(* Logix 5000 project; controller FV vendor 1 type 14 code 217 rev 31.11; software revision 31.00; part 47 of 63 *)
(* tags used below, declared in another part *)
   CWD : CHECKWORD_FLAGS;
   Delphi_Does_Eng_Func : BOOL;
   FV_FV13C : PlantItem;   // FV13C
   FV_FV13J : PlantItem;   // FV13J
   FV_FV14C : PlantItem;   // FV14C
   FV_FV14J : PlantItem;   // FV14J
   FV_FV15C : PlantItem;   // FV15C
   FV_FV15J : PlantItem;   // FV15J
   FV_FV16C : PlantItem;   // FV16C
   FV_FV16J : PlantItem;   // FV16J
   FV_FV17C : PlantItem;   // FV17C
   FV_FV17J : PlantItem;   // FV17J
   FV_FV18C : PlantItem;   // FV18C
   FV_FV18J : PlantItem;   // FV18J
   FV_FV19C : PlantItem;   // FV19C
   FV_FV19J : PlantItem;   // FV19J
   FV_FV20C : PlantItem;   // FV20C
   FV_FV20J : PlantItem;   // FV20J
   FV_FV21C : PlantItem;   // FV21C
   FV_FV21J : PlantItem;   // FV21J
   FV_FV22C : PlantItem;   // FV22C
   FV_FV22J : PlantItem;   // FV22J
   FV_FV23C : PlantItem;   // FV23C
   FV_FV23J : PlantItem;   // FV23J
   FV_FV24C : PlantItem;   // FV24C
   FV_FV24J : PlantItem;   // FV24J
   FV_N255 : INT[255];   // Old Checkwords to keep Delphi working in the interim before full changeover.
(* FV_Common, continued *)

   24: [XIC(Delphi_Does_Eng_Func) [[XIC(FV_N255[25].8) [OTL(FV_FV13C.CW.[CWD.MANUAL]) ,XIC(FV_N255[25].9) OTL(FV_FV13C.CW.[CWD.MANDRV]) ,XIO(FV_N255[25].9) OTU(FV_FV13C.CW.[CWD.MANDRV]) ] ,XIO(FV_N255[25].8) [OTU(FV_FV13C.CW.[CWD.MANUAL]) ,[XIC(FV_FV13C.CW.[CWD.OUTPUT]) OTL(FV_N255[25].9) ,XIO(FV_FV13C.CW.[CWD.OUTPUT]) OTU(FV_N255[25].9) ] ] ] ,[XIC(FV_N255[25].13) OTL(FV_FV13C.CW.[CWD.CHECKOFF]) ,XIO(FV_N255[25].13) OTU(FV_FV13C.CW.[CWD.CHECKOFF]) ] ] ,XIO(Delphi_Does_Eng_Func) [[XIC(FV_FV13C.CW.[CWD.MANUAL]) OTL(FV_N255[25].8) ,XIO(FV_FV13C.CW.[CWD.MANUAL]) OTU(FV_N255[25].8) ] ,[XIC(FV_FV13C.CW.[CWD.CHECKOFF]) OTL(FV_N255[25].13) ,XIO(FV_FV13C.CW.[CWD.CHECKOFF]) OTU(FV_N255[25].13) ] ,[XIC(FV_FV13C.CW.[CWD.OUTPUT]) OTL(FV_N255[25].9) ,XIO(FV_FV13C.CW.[CWD.OUTPUT]) OTU(FV_N255[25].9) ] ] ,XIC(FV_FV13C.CW.[CWD.OUTPUT]) OTE(FV_N255[25].10) ,XIO(FV_FV13C.CW.[CWD.OUTPUT]) OTE(FV_N255[25].11) ,XIC(FV_FV13C.CW.[CWD.FAULT]) OTE(FV_N255[25].15) ];
   25: [XIC(Delphi_Does_Eng_Func) [[XIC(FV_N255[26].8) [OTL(FV_FV13J.CW.[CWD.MANUAL]) ,XIC(FV_N255[26].9) OTL(FV_FV13J.CW.[CWD.MANDRV]) ,XIO(FV_N255[26].9) OTU(FV_FV13J.CW.[CWD.MANDRV]) ] ,XIO(FV_N255[26].8) [OTU(FV_FV13J.CW.[CWD.MANUAL]) ,[XIC(FV_FV13J.CW.[CWD.OUTPUT]) OTL(FV_N255[26].9) ,XIO(FV_FV13J.CW.[CWD.OUTPUT]) OTU(FV_N255[26].9) ] ] ] ,[XIC(FV_N255[26].13) OTL(FV_FV13J.CW.[CWD.CHECKOFF]) ,XIO(FV_N255[26].13) OTU(FV_FV13J.CW.[CWD.CHECKOFF]) ] ] ,XIO(Delphi_Does_Eng_Func) [[XIC(FV_FV13J.CW.[CWD.MANUAL]) OTL(FV_N255[26].8) ,XIO(FV_FV13J.CW.[CWD.MANUAL]) OTU(FV_N255[26].8) ] ,[XIC(FV_FV13J.CW.[CWD.CHECKOFF]) OTL(FV_N255[26].13) ,XIO(FV_FV13J.CW.[CWD.CHECKOFF]) OTU(FV_N255[26].13) ] ,[XIC(FV_FV13J.CW.[CWD.OUTPUT]) OTL(FV_N255[26].9) ,XIO(FV_FV13J.CW.[CWD.OUTPUT]) OTU(FV_N255[26].9) ] ] ,XIC(FV_FV13J.CW.[CWD.OUTPUT]) OTE(FV_N255[26].10) ,XIO(FV_FV13J.CW.[CWD.OUTPUT]) OTE(FV_N255[26].11) ,XIC(FV_FV13J.CW.[CWD.FAULT]) OTE(FV_N255[26].15) ];
   26: [XIC(Delphi_Does_Eng_Func) [[XIC(FV_N255[27].8) [OTL(FV_FV14C.CW.[CWD.MANUAL]) ,XIC(FV_N255[27].9) OTL(FV_FV14C.CW.[CWD.MANDRV]) ,XIO(FV_N255[27].9) OTU(FV_FV14C.CW.[CWD.MANDRV]) ] ,XIO(FV_N255[27].8) [OTU(FV_FV14C.CW.[CWD.MANUAL]) ,[XIC(FV_FV14C.CW.[CWD.OUTPUT]) OTL(FV_N255[27].9) ,XIO(FV_FV14C.CW.[CWD.OUTPUT]) OTU(FV_N255[27].9) ] ] ] ,[XIC(FV_N255[27].13) OTL(FV_FV14C.CW.[CWD.CHECKOFF]) ,XIO(FV_N255[27].13) OTU(FV_FV14C.CW.[CWD.CHECKOFF]) ] ] ,XIO(Delphi_Does_Eng_Func) [[XIC(FV_FV14C.CW.[CWD.MANUAL]) OTL(FV_N255[27].8) ,XIO(FV_FV14C.CW.[CWD.MANUAL]) OTU(FV_N255[27].8) ] ,[XIC(FV_FV14C.CW.[CWD.CHECKOFF]) OTL(FV_N255[27].13) ,XIO(FV_FV14C.CW.[CWD.CHECKOFF]) OTU(FV_N255[27].13) ] ,[XIC(FV_FV14C.CW.[CWD.OUTPUT]) OTL(FV_N255[27].9) ,XIO(FV_FV14C.CW.[CWD.OUTPUT]) OTU(FV_N255[27].9) ] ] ,XIC(FV_FV14C.CW.[CWD.OUTPUT]) OTE(FV_N255[27].10) ,XIO(FV_FV14C.CW.[CWD.OUTPUT]) OTE(FV_N255[27].11) ,XIC(FV_FV14C.CW.[CWD.FAULT]) OTE(FV_N255[27].15) ];
   27: [XIC(Delphi_Does_Eng_Func) [[XIC(FV_N255[28].8) [OTL(FV_FV14J.CW.[CWD.MANUAL]) ,XIC(FV_N255[28].9) OTL(FV_FV14J.CW.[CWD.MANDRV]) ,XIO(FV_N255[28].9) OTU(FV_FV14J.CW.[CWD.MANDRV]) ] ,XIO(FV_N255[28].8) [OTU(FV_FV14J.CW.[CWD.MANUAL]) ,[XIC(FV_FV14J.CW.[CWD.OUTPUT]) OTL(FV_N255[28].9) ,XIO(FV_FV14J.CW.[CWD.OUTPUT]) OTU(FV_N255[28].9) ] ] ] ,[XIC(FV_N255[28].13) OTL(FV_FV14J.CW.[CWD.CHECKOFF]) ,XIO(FV_N255[28].13) OTU(FV_FV14J.CW.[CWD.CHECKOFF]) ] ] ,XIO(Delphi_Does_Eng_Func) [[XIC(FV_FV14J.CW.[CWD.MANUAL]) OTL(FV_N255[28].8) ,XIO(FV_FV14J.CW.[CWD.MANUAL]) OTU(FV_N255[28].8) ] ,[XIC(FV_FV14J.CW.[CWD.CHECKOFF]) OTL(FV_N255[28].13) ,XIO(FV_FV14J.CW.[CWD.CHECKOFF]) OTU(FV_N255[28].13) ] ,[XIC(FV_FV14J.CW.[CWD.OUTPUT]) OTL(FV_N255[28].9) ,XIO(FV_FV14J.CW.[CWD.OUTPUT]) OTU(FV_N255[28].9) ] ] ,XIC(FV_FV14J.CW.[CWD.OUTPUT]) OTE(FV_N255[28].10) ,XIO(FV_FV14J.CW.[CWD.OUTPUT]) OTE(FV_N255[28].11) ,XIC(FV_FV14J.CW.[CWD.FAULT]) OTE(FV_N255[28].15) ];
   28: [XIC(Delphi_Does_Eng_Func) [[XIC(FV_N255[29].8) [OTL(FV_FV15C.CW.[CWD.MANUAL]) ,XIC(FV_N255[29].9) OTL(FV_FV15C.CW.[CWD.MANDRV]) ,XIO(FV_N255[29].9) OTU(FV_FV15C.CW.[CWD.MANDRV]) ] ,XIO(FV_N255[29].8) [OTU(FV_FV15C.CW.[CWD.MANUAL]) ,[XIC(FV_FV15C.CW.[CWD.OUTPUT]) OTL(FV_N255[29].9) ,XIO(FV_FV15C.CW.[CWD.OUTPUT]) OTU(FV_N255[29].9) ] ] ] ,[XIC(FV_N255[29].13) OTL(FV_FV15C.CW.[CWD.CHECKOFF]) ,XIO(FV_N255[29].13) OTU(FV_FV15C.CW.[CWD.CHECKOFF]) ] ] ,XIO(Delphi_Does_Eng_Func) [[XIC(FV_FV15C.CW.[CWD.MANUAL]) OTL(FV_N255[29].8) ,XIO(FV_FV15C.CW.[CWD.MANUAL]) OTU(FV_N255[29].8) ] ,[XIC(FV_FV15C.CW.[CWD.CHECKOFF]) OTL(FV_N255[29].13) ,XIO(FV_FV15C.CW.[CWD.CHECKOFF]) OTU(FV_N255[29].13) ] ,[XIC(FV_FV15C.CW.[CWD.OUTPUT]) OTL(FV_N255[29].9) ,XIO(FV_FV15C.CW.[CWD.OUTPUT]) OTU(FV_N255[29].9) ] ] ,XIC(FV_FV15C.CW.[CWD.OUTPUT]) OTE(FV_N255[29].10) ,XIO(FV_FV15C.CW.[CWD.OUTPUT]) OTE(FV_N255[29].11) ,XIC(FV_FV15C.CW.[CWD.FAULT]) OTE(FV_N255[29].15) ];
   29: [XIC(Delphi_Does_Eng_Func) [[XIC(FV_N255[30].8) [OTL(FV_FV15J.CW.[CWD.MANUAL]) ,XIC(FV_N255[30].9) OTL(FV_FV15J.CW.[CWD.MANDRV]) ,XIO(FV_N255[30].9) OTU(FV_FV15J.CW.[CWD.MANDRV]) ] ,XIO(FV_N255[30].8) [OTU(FV_FV15J.CW.[CWD.MANUAL]) ,[XIC(FV_FV15J.CW.[CWD.OUTPUT]) OTL(FV_N255[30].9) ,XIO(FV_FV15J.CW.[CWD.OUTPUT]) OTU(FV_N255[30].9) ] ] ] ,[XIC(FV_N255[30].13) OTL(FV_FV15J.CW.[CWD.CHECKOFF]) ,XIO(FV_N255[30].13) OTU(FV_FV15J.CW.[CWD.CHECKOFF]) ] ] ,XIO(Delphi_Does_Eng_Func) [[XIC(FV_FV15J.CW.[CWD.MANUAL]) OTL(FV_N255[30].8) ,XIO(FV_FV15J.CW.[CWD.MANUAL]) OTU(FV_N255[30].8) ] ,[XIC(FV_FV15J.CW.[CWD.CHECKOFF]) OTL(FV_N255[30].13) ,XIO(FV_FV15J.CW.[CWD.CHECKOFF]) OTU(FV_N255[30].13) ] ,[XIC(FV_FV15J.CW.[CWD.OUTPUT]) OTL(FV_N255[30].9) ,XIO(FV_FV15J.CW.[CWD.OUTPUT]) OTU(FV_N255[30].9) ] ] ,XIC(FV_FV15J.CW.[CWD.OUTPUT]) OTE(FV_N255[30].10) ,XIO(FV_FV15J.CW.[CWD.OUTPUT]) OTE(FV_N255[30].11) ,XIC(FV_FV15J.CW.[CWD.FAULT]) OTE(FV_N255[30].15) ];
   30: [XIC(Delphi_Does_Eng_Func) [[XIC(FV_N255[31].8) [OTL(FV_FV16C.CW.[CWD.MANUAL]) ,XIC(FV_N255[31].9) OTL(FV_FV16C.CW.[CWD.MANDRV]) ,XIO(FV_N255[31].9) OTU(FV_FV16C.CW.[CWD.MANDRV]) ] ,XIO(FV_N255[31].8) [OTU(FV_FV16C.CW.[CWD.MANUAL]) ,[XIC(FV_FV16C.CW.[CWD.OUTPUT]) OTL(FV_N255[31].9) ,XIO(FV_FV16C.CW.[CWD.OUTPUT]) OTU(FV_N255[31].9) ] ] ] ,[XIC(FV_N255[31].13) OTL(FV_FV16C.CW.[CWD.CHECKOFF]) ,XIO(FV_N255[31].13) OTU(FV_FV16C.CW.[CWD.CHECKOFF]) ] ] ,XIO(Delphi_Does_Eng_Func) [[XIC(FV_FV16C.CW.[CWD.MANUAL]) OTL(FV_N255[31].8) ,XIO(FV_FV16C.CW.[CWD.MANUAL]) OTU(FV_N255[31].8) ] ,[XIC(FV_FV16C.CW.[CWD.CHECKOFF]) OTL(FV_N255[31].13) ,XIO(FV_FV16C.CW.[CWD.CHECKOFF]) OTU(FV_N255[31].13) ] ,[XIC(FV_FV16C.CW.[CWD.OUTPUT]) OTL(FV_N255[31].9) ,XIO(FV_FV16C.CW.[CWD.OUTPUT]) OTU(FV_N255[31].9) ] ] ,XIC(FV_FV16C.CW.[CWD.OUTPUT]) OTE(FV_N255[31].10) ,XIO(FV_FV16C.CW.[CWD.OUTPUT]) OTE(FV_N255[31].11) ,XIC(FV_FV16C.CW.[CWD.FAULT]) OTE(FV_N255[31].15) ];
   31: [XIC(Delphi_Does_Eng_Func) [[XIC(FV_N255[32].8) [OTL(FV_FV16J.CW.[CWD.MANUAL]) ,XIC(FV_N255[32].9) OTL(FV_FV16J.CW.[CWD.MANDRV]) ,XIO(FV_N255[32].9) OTU(FV_FV16J.CW.[CWD.MANDRV]) ] ,XIO(FV_N255[32].8) [OTU(FV_FV16J.CW.[CWD.MANUAL]) ,[XIC(FV_FV16J.CW.[CWD.OUTPUT]) OTL(FV_N255[32].9) ,XIO(FV_FV16J.CW.[CWD.OUTPUT]) OTU(FV_N255[32].9) ] ] ] ,[XIC(FV_N255[32].13) OTL(FV_FV16J.CW.[CWD.CHECKOFF]) ,XIO(FV_N255[32].13) OTU(FV_FV16J.CW.[CWD.CHECKOFF]) ] ] ,XIO(Delphi_Does_Eng_Func) [[XIC(FV_FV16J.CW.[CWD.MANUAL]) OTL(FV_N255[32].8) ,XIO(FV_FV16J.CW.[CWD.MANUAL]) OTU(FV_N255[32].8) ] ,[XIC(FV_FV16J.CW.[CWD.CHECKOFF]) OTL(FV_N255[32].13) ,XIO(FV_FV16J.CW.[CWD.CHECKOFF]) OTU(FV_N255[32].13) ] ,[XIC(FV_FV16J.CW.[CWD.OUTPUT]) OTL(FV_N255[32].9) ,XIO(FV_FV16J.CW.[CWD.OUTPUT]) OTU(FV_N255[32].9) ] ] ,XIC(FV_FV16J.CW.[CWD.OUTPUT]) OTE(FV_N255[32].10) ,XIO(FV_FV16J.CW.[CWD.OUTPUT]) OTE(FV_N255[32].11) ,XIC(FV_FV16J.CW.[CWD.FAULT]) OTE(FV_N255[32].15) ];
   32: [XIC(Delphi_Does_Eng_Func) [[XIC(FV_N255[33].8) [OTL(FV_FV17C.CW.[CWD.MANUAL]) ,XIC(FV_N255[33].9) OTL(FV_FV17C.CW.[CWD.MANDRV]) ,XIO(FV_N255[33].9) OTU(FV_FV17C.CW.[CWD.MANDRV]) ] ,XIO(FV_N255[33].8) [OTU(FV_FV17C.CW.[CWD.MANUAL]) ,[XIC(FV_FV17C.CW.[CWD.OUTPUT]) OTL(FV_N255[33].9) ,XIO(FV_FV17C.CW.[CWD.OUTPUT]) OTU(FV_N255[33].9) ] ] ] ,[XIC(FV_N255[33].13) OTL(FV_FV17C.CW.[CWD.CHECKOFF]) ,XIO(FV_N255[33].13) OTU(FV_FV17C.CW.[CWD.CHECKOFF]) ] ] ,XIO(Delphi_Does_Eng_Func) [[XIC(FV_FV17C.CW.[CWD.MANUAL]) OTL(FV_N255[33].8) ,XIO(FV_FV17C.CW.[CWD.MANUAL]) OTU(FV_N255[33].8) ] ,[XIC(FV_FV17C.CW.[CWD.CHECKOFF]) OTL(FV_N255[33].13) ,XIO(FV_FV17C.CW.[CWD.CHECKOFF]) OTU(FV_N255[33].13) ] ,[XIC(FV_FV17C.CW.[CWD.OUTPUT]) OTL(FV_N255[33].9) ,XIO(FV_FV17C.CW.[CWD.OUTPUT]) OTU(FV_N255[33].9) ] ] ,XIC(FV_FV17C.CW.[CWD.OUTPUT]) OTE(FV_N255[33].10) ,XIO(FV_FV17C.CW.[CWD.OUTPUT]) OTE(FV_N255[33].11) ,XIC(FV_FV17C.CW.[CWD.FAULT]) OTE(FV_N255[33].15) ];
   33: [XIC(Delphi_Does_Eng_Func) [[XIC(FV_N255[34].8) [OTL(FV_FV17J.CW.[CWD.MANUAL]) ,XIC(FV_N255[34].9) OTL(FV_FV17J.CW.[CWD.MANDRV]) ,XIO(FV_N255[34].9) OTU(FV_FV17J.CW.[CWD.MANDRV]) ] ,XIO(FV_N255[34].8) [OTU(FV_FV17J.CW.[CWD.MANUAL]) ,[XIC(FV_FV17J.CW.[CWD.OUTPUT]) OTL(FV_N255[34].9) ,XIO(FV_FV17J.CW.[CWD.OUTPUT]) OTU(FV_N255[34].9) ] ] ] ,[XIC(FV_N255[34].13) OTL(FV_FV17J.CW.[CWD.CHECKOFF]) ,XIO(FV_N255[34].13) OTU(FV_FV17J.CW.[CWD.CHECKOFF]) ] ] ,XIO(Delphi_Does_Eng_Func) [[XIC(FV_FV17J.CW.[CWD.MANUAL]) OTL(FV_N255[34].8) ,XIO(FV_FV17J.CW.[CWD.MANUAL]) OTU(FV_N255[34].8) ] ,[XIC(FV_FV17J.CW.[CWD.CHECKOFF]) OTL(FV_N255[34].13) ,XIO(FV_FV17J.CW.[CWD.CHECKOFF]) OTU(FV_N255[34].13) ] ,[XIC(FV_FV17J.CW.[CWD.OUTPUT]) OTL(FV_N255[34].9) ,XIO(FV_FV17J.CW.[CWD.OUTPUT]) OTU(FV_N255[34].9) ] ] ,XIC(FV_FV17J.CW.[CWD.OUTPUT]) OTE(FV_N255[34].10) ,XIO(FV_FV17J.CW.[CWD.OUTPUT]) OTE(FV_N255[34].11) ,XIC(FV_FV17J.CW.[CWD.FAULT]) OTE(FV_N255[34].15) ];
   34: [XIC(Delphi_Does_Eng_Func) [[XIC(FV_N255[35].8) [OTL(FV_FV18C.CW.[CWD.MANUAL]) ,XIC(FV_N255[35].9) OTL(FV_FV18C.CW.[CWD.MANDRV]) ,XIO(FV_N255[35].9) OTU(FV_FV18C.CW.[CWD.MANDRV]) ] ,XIO(FV_N255[35].8) [OTU(FV_FV18C.CW.[CWD.MANUAL]) ,[XIC(FV_FV18C.CW.[CWD.OUTPUT]) OTL(FV_N255[35].9) ,XIO(FV_FV18C.CW.[CWD.OUTPUT]) OTU(FV_N255[35].9) ] ] ] ,[XIC(FV_N255[35].13) OTL(FV_FV18C.CW.[CWD.CHECKOFF]) ,XIO(FV_N255[35].13) OTU(FV_FV18C.CW.[CWD.CHECKOFF]) ] ] ,XIO(Delphi_Does_Eng_Func) [[XIC(FV_FV18C.CW.[CWD.MANUAL]) OTL(FV_N255[35].8) ,XIO(FV_FV18C.CW.[CWD.MANUAL]) OTU(FV_N255[35].8) ] ,[XIC(FV_FV18C.CW.[CWD.CHECKOFF]) OTL(FV_N255[35].13) ,XIO(FV_FV18C.CW.[CWD.CHECKOFF]) OTU(FV_N255[35].13) ] ,[XIC(FV_FV18C.CW.[CWD.OUTPUT]) OTL(FV_N255[35].9) ,XIO(FV_FV18C.CW.[CWD.OUTPUT]) OTU(FV_N255[35].9) ] ] ,XIC(FV_FV18C.CW.[CWD.OUTPUT]) OTE(FV_N255[35].10) ,XIO(FV_FV18C.CW.[CWD.OUTPUT]) OTE(FV_N255[35].11) ,XIC(FV_FV18C.CW.[CWD.FAULT]) OTE(FV_N255[35].15) ];
   35: [XIC(Delphi_Does_Eng_Func) [[XIC(FV_N255[36].8) [OTL(FV_FV18J.CW.[CWD.MANUAL]) ,XIC(FV_N255[36].9) OTL(FV_FV18J.CW.[CWD.MANDRV]) ,XIO(FV_N255[36].9) OTU(FV_FV18J.CW.[CWD.MANDRV]) ] ,XIO(FV_N255[36].8) [OTU(FV_FV18J.CW.[CWD.MANUAL]) ,[XIC(FV_FV18J.CW.[CWD.OUTPUT]) OTL(FV_N255[36].9) ,XIO(FV_FV18J.CW.[CWD.OUTPUT]) OTU(FV_N255[36].9) ] ] ] ,[XIC(FV_N255[36].13) OTL(FV_FV18J.CW.[CWD.CHECKOFF]) ,XIO(FV_N255[36].13) OTU(FV_FV18J.CW.[CWD.CHECKOFF]) ] ] ,XIO(Delphi_Does_Eng_Func) [[XIC(FV_FV18J.CW.[CWD.MANUAL]) OTL(FV_N255[36].8) ,XIO(FV_FV18J.CW.[CWD.MANUAL]) OTU(FV_N255[36].8) ] ,[XIC(FV_FV18J.CW.[CWD.CHECKOFF]) OTL(FV_N255[36].13) ,XIO(FV_FV18J.CW.[CWD.CHECKOFF]) OTU(FV_N255[36].13) ] ,[XIC(FV_FV18J.CW.[CWD.OUTPUT]) OTL(FV_N255[36].9) ,XIO(FV_FV18J.CW.[CWD.OUTPUT]) OTU(FV_N255[36].9) ] ] ,XIC(FV_FV18J.CW.[CWD.OUTPUT]) OTE(FV_N255[36].10) ,XIO(FV_FV18J.CW.[CWD.OUTPUT]) OTE(FV_N255[36].11) ,XIC(FV_FV18J.CW.[CWD.FAULT]) OTE(FV_N255[36].15) ];
   36: [XIC(Delphi_Does_Eng_Func) [[XIC(FV_N255[37].8) [OTL(FV_FV19C.CW.[CWD.MANUAL]) ,XIC(FV_N255[37].9) OTL(FV_FV19C.CW.[CWD.MANDRV]) ,XIO(FV_N255[37].9) OTU(FV_FV19C.CW.[CWD.MANDRV]) ] ,XIO(FV_N255[37].8) [OTU(FV_FV19C.CW.[CWD.MANUAL]) ,[XIC(FV_FV19C.CW.[CWD.OUTPUT]) OTL(FV_N255[37].9) ,XIO(FV_FV19C.CW.[CWD.OUTPUT]) OTU(FV_N255[37].9) ] ] ] ,[XIC(FV_N255[37].13) OTL(FV_FV19C.CW.[CWD.CHECKOFF]) ,XIO(FV_N255[37].13) OTU(FV_FV19C.CW.[CWD.CHECKOFF]) ] ] ,XIO(Delphi_Does_Eng_Func) [[XIC(FV_FV19C.CW.[CWD.MANUAL]) OTL(FV_N255[37].8) ,XIO(FV_FV19C.CW.[CWD.MANUAL]) OTU(FV_N255[37].8) ] ,[XIC(FV_FV19C.CW.[CWD.CHECKOFF]) OTL(FV_N255[37].13) ,XIO(FV_FV19C.CW.[CWD.CHECKOFF]) OTU(FV_N255[37].13) ] ,[XIC(FV_FV19C.CW.[CWD.OUTPUT]) OTL(FV_N255[37].9) ,XIO(FV_FV19C.CW.[CWD.OUTPUT]) OTU(FV_N255[37].9) ] ] ,XIC(FV_FV19C.CW.[CWD.OUTPUT]) OTE(FV_N255[37].10) ,XIO(FV_FV19C.CW.[CWD.OUTPUT]) OTE(FV_N255[37].11) ,XIC(FV_FV19C.CW.[CWD.FAULT]) OTE(FV_N255[37].15) ];
   37: [XIC(Delphi_Does_Eng_Func) [[XIC(FV_N255[38].8) [OTL(FV_FV19J.CW.[CWD.MANUAL]) ,XIC(FV_N255[38].9) OTL(FV_FV19J.CW.[CWD.MANDRV]) ,XIO(FV_N255[38].9) OTU(FV_FV19J.CW.[CWD.MANDRV]) ] ,XIO(FV_N255[38].8) [OTU(FV_FV19J.CW.[CWD.MANUAL]) ,[XIC(FV_FV19J.CW.[CWD.OUTPUT]) OTL(FV_N255[38].9) ,XIO(FV_FV19J.CW.[CWD.OUTPUT]) OTU(FV_N255[38].9) ] ] ] ,[XIC(FV_N255[38].13) OTL(FV_FV19J.CW.[CWD.CHECKOFF]) ,XIO(FV_N255[38].13) OTU(FV_FV19J.CW.[CWD.CHECKOFF]) ] ] ,XIO(Delphi_Does_Eng_Func) [[XIC(FV_FV19J.CW.[CWD.MANUAL]) OTL(FV_N255[38].8) ,XIO(FV_FV19J.CW.[CWD.MANUAL]) OTU(FV_N255[38].8) ] ,[XIC(FV_FV19J.CW.[CWD.CHECKOFF]) OTL(FV_N255[38].13) ,XIO(FV_FV19J.CW.[CWD.CHECKOFF]) OTU(FV_N255[38].13) ] ,[XIC(FV_FV19J.CW.[CWD.OUTPUT]) OTL(FV_N255[38].9) ,XIO(FV_FV19J.CW.[CWD.OUTPUT]) OTU(FV_N255[38].9) ] ] ,XIC(FV_FV19J.CW.[CWD.OUTPUT]) OTE(FV_N255[38].10) ,XIO(FV_FV19J.CW.[CWD.OUTPUT]) OTE(FV_N255[38].11) ,XIC(FV_FV19J.CW.[CWD.FAULT]) OTE(FV_N255[38].15) ];
   38: [XIC(Delphi_Does_Eng_Func) [[XIC(FV_N255[39].8) [OTL(FV_FV20C.CW.[CWD.MANUAL]) ,XIC(FV_N255[39].9) OTL(FV_FV20C.CW.[CWD.MANDRV]) ,XIO(FV_N255[39].9) OTU(FV_FV20C.CW.[CWD.MANDRV]) ] ,XIO(FV_N255[39].8) [OTU(FV_FV20C.CW.[CWD.MANUAL]) ,[XIC(FV_FV20C.CW.[CWD.OUTPUT]) OTL(FV_N255[39].9) ,XIO(FV_FV20C.CW.[CWD.OUTPUT]) OTU(FV_N255[39].9) ] ] ] ,[XIC(FV_N255[39].13) OTL(FV_FV20C.CW.[CWD.CHECKOFF]) ,XIO(FV_N255[39].13) OTU(FV_FV20C.CW.[CWD.CHECKOFF]) ] ] ,XIO(Delphi_Does_Eng_Func) [[XIC(FV_FV20C.CW.[CWD.MANUAL]) OTL(FV_N255[39].8) ,XIO(FV_FV20C.CW.[CWD.MANUAL]) OTU(FV_N255[39].8) ] ,[XIC(FV_FV20C.CW.[CWD.CHECKOFF]) OTL(FV_N255[39].13) ,XIO(FV_FV20C.CW.[CWD.CHECKOFF]) OTU(FV_N255[39].13) ] ,[XIC(FV_FV20C.CW.[CWD.OUTPUT]) OTL(FV_N255[39].9) ,XIO(FV_FV20C.CW.[CWD.OUTPUT]) OTU(FV_N255[39].9) ] ] ,XIC(FV_FV20C.CW.[CWD.OUTPUT]) OTE(FV_N255[39].10) ,XIO(FV_FV20C.CW.[CWD.OUTPUT]) OTE(FV_N255[39].11) ,XIC(FV_FV20C.CW.[CWD.FAULT]) OTE(FV_N255[39].15) ];
   39: [XIC(Delphi_Does_Eng_Func) [[XIC(FV_N255[40].8) [OTL(FV_FV20J.CW.[CWD.MANUAL]) ,XIC(FV_N255[40].9) OTL(FV_FV20J.CW.[CWD.MANDRV]) ,XIO(FV_N255[40].9) OTU(FV_FV20J.CW.[CWD.MANDRV]) ] ,XIO(FV_N255[40].8) [OTU(FV_FV20J.CW.[CWD.MANUAL]) ,[XIC(FV_FV20J.CW.[CWD.OUTPUT]) OTL(FV_N255[40].9) ,XIO(FV_FV20J.CW.[CWD.OUTPUT]) OTU(FV_N255[40].9) ] ] ] ,[XIC(FV_N255[40].13) OTL(FV_FV20J.CW.[CWD.CHECKOFF]) ,XIO(FV_N255[40].13) OTU(FV_FV20J.CW.[CWD.CHECKOFF]) ] ] ,XIO(Delphi_Does_Eng_Func) [[XIC(FV_FV20J.CW.[CWD.MANUAL]) OTL(FV_N255[40].8) ,XIO(FV_FV20J.CW.[CWD.MANUAL]) OTU(FV_N255[40].8) ] ,[XIC(FV_FV20J.CW.[CWD.CHECKOFF]) OTL(FV_N255[40].13) ,XIO(FV_FV20J.CW.[CWD.CHECKOFF]) OTU(FV_N255[40].13) ] ,[XIC(FV_FV20J.CW.[CWD.OUTPUT]) OTL(FV_N255[40].9) ,XIO(FV_FV20J.CW.[CWD.OUTPUT]) OTU(FV_N255[40].9) ] ] ,XIC(FV_FV20J.CW.[CWD.OUTPUT]) OTE(FV_N255[40].10) ,XIO(FV_FV20J.CW.[CWD.OUTPUT]) OTE(FV_N255[40].11) ,XIC(FV_FV20J.CW.[CWD.FAULT]) OTE(FV_N255[40].15) ];
   40: [XIC(Delphi_Does_Eng_Func) [[XIC(FV_N255[41].8) [OTL(FV_FV21C.CW.[CWD.MANUAL]) ,XIC(FV_N255[41].9) OTL(FV_FV21C.CW.[CWD.MANDRV]) ,XIO(FV_N255[41].9) OTU(FV_FV21C.CW.[CWD.MANDRV]) ] ,XIO(FV_N255[41].8) [OTU(FV_FV21C.CW.[CWD.MANUAL]) ,[XIC(FV_FV21C.CW.[CWD.OUTPUT]) OTL(FV_N255[41].9) ,XIO(FV_FV21C.CW.[CWD.OUTPUT]) OTU(FV_N255[41].9) ] ] ] ,[XIC(FV_N255[41].13) OTL(FV_FV21C.CW.[CWD.CHECKOFF]) ,XIO(FV_N255[41].13) OTU(FV_FV21C.CW.[CWD.CHECKOFF]) ] ] ,XIO(Delphi_Does_Eng_Func) [[XIC(FV_FV21C.CW.[CWD.MANUAL]) OTL(FV_N255[41].8) ,XIO(FV_FV21C.CW.[CWD.MANUAL]) OTU(FV_N255[41].8) ] ,[XIC(FV_FV21C.CW.[CWD.CHECKOFF]) OTL(FV_N255[41].13) ,XIO(FV_FV21C.CW.[CWD.CHECKOFF]) OTU(FV_N255[41].13) ] ,[XIC(FV_FV21C.CW.[CWD.OUTPUT]) OTL(FV_N255[41].9) ,XIO(FV_FV21C.CW.[CWD.OUTPUT]) OTU(FV_N255[41].9) ] ] ,XIC(FV_FV21C.CW.[CWD.OUTPUT]) OTE(FV_N255[41].10) ,XIO(FV_FV21C.CW.[CWD.OUTPUT]) OTE(FV_N255[41].11) ,XIC(FV_FV21C.CW.[CWD.FAULT]) OTE(FV_N255[41].15) ];
   41: [XIC(Delphi_Does_Eng_Func) [[XIC(FV_N255[42].8) [OTL(FV_FV21J.CW.[CWD.MANUAL]) ,XIC(FV_N255[42].9) OTL(FV_FV21J.CW.[CWD.MANDRV]) ,XIO(FV_N255[42].9) OTU(FV_FV21J.CW.[CWD.MANDRV]) ] ,XIO(FV_N255[42].8) [OTU(FV_FV21J.CW.[CWD.MANUAL]) ,[XIC(FV_FV21J.CW.[CWD.OUTPUT]) OTL(FV_N255[42].9) ,XIO(FV_FV21J.CW.[CWD.OUTPUT]) OTU(FV_N255[42].9) ] ] ] ,[XIC(FV_N255[42].13) OTL(FV_FV21J.CW.[CWD.CHECKOFF]) ,XIO(FV_N255[42].13) OTU(FV_FV21J.CW.[CWD.CHECKOFF]) ] ] ,XIO(Delphi_Does_Eng_Func) [[XIC(FV_FV21J.CW.[CWD.MANUAL]) OTL(FV_N255[42].8) ,XIO(FV_FV21J.CW.[CWD.MANUAL]) OTU(FV_N255[42].8) ] ,[XIC(FV_FV21J.CW.[CWD.CHECKOFF]) OTL(FV_N255[42].13) ,XIO(FV_FV21J.CW.[CWD.CHECKOFF]) OTU(FV_N255[42].13) ] ,[XIC(FV_FV21J.CW.[CWD.OUTPUT]) OTL(FV_N255[42].9) ,XIO(FV_FV21J.CW.[CWD.OUTPUT]) OTU(FV_N255[42].9) ] ] ,XIC(FV_FV21J.CW.[CWD.OUTPUT]) OTE(FV_N255[42].10) ,XIO(FV_FV21J.CW.[CWD.OUTPUT]) OTE(FV_N255[42].11) ,XIC(FV_FV21J.CW.[CWD.FAULT]) OTE(FV_N255[42].15) ];
   42: [XIC(Delphi_Does_Eng_Func) [[XIC(FV_N255[43].8) [OTL(FV_FV22C.CW.[CWD.MANUAL]) ,XIC(FV_N255[43].9) OTL(FV_FV22C.CW.[CWD.MANDRV]) ,XIO(FV_N255[43].9) OTU(FV_FV22C.CW.[CWD.MANDRV]) ] ,XIO(FV_N255[43].8) [OTU(FV_FV22C.CW.[CWD.MANUAL]) ,[XIC(FV_FV22C.CW.[CWD.OUTPUT]) OTL(FV_N255[43].9) ,XIO(FV_FV22C.CW.[CWD.OUTPUT]) OTU(FV_N255[43].9) ] ] ] ,[XIC(FV_N255[43].13) OTL(FV_FV22C.CW.[CWD.CHECKOFF]) ,XIO(FV_N255[43].13) OTU(FV_FV22C.CW.[CWD.CHECKOFF]) ] ] ,XIO(Delphi_Does_Eng_Func) [[XIC(FV_FV22C.CW.[CWD.MANUAL]) OTL(FV_N255[43].8) ,XIO(FV_FV22C.CW.[CWD.MANUAL]) OTU(FV_N255[43].8) ] ,[XIC(FV_FV22C.CW.[CWD.CHECKOFF]) OTL(FV_N255[43].13) ,XIO(FV_FV22C.CW.[CWD.CHECKOFF]) OTU(FV_N255[43].13) ] ,[XIC(FV_FV22C.CW.[CWD.OUTPUT]) OTL(FV_N255[43].9) ,XIO(FV_FV22C.CW.[CWD.OUTPUT]) OTU(FV_N255[43].9) ] ] ,XIC(FV_FV22C.CW.[CWD.OUTPUT]) OTE(FV_N255[43].10) ,XIO(FV_FV22C.CW.[CWD.OUTPUT]) OTE(FV_N255[43].11) ,XIC(FV_FV22C.CW.[CWD.FAULT]) OTE(FV_N255[43].15) ];
   43: [XIC(Delphi_Does_Eng_Func) [[XIC(FV_N255[44].8) [OTL(FV_FV22J.CW.[CWD.MANUAL]) ,XIC(FV_N255[44].9) OTL(FV_FV22J.CW.[CWD.MANDRV]) ,XIO(FV_N255[44].9) OTU(FV_FV22J.CW.[CWD.MANDRV]) ] ,XIO(FV_N255[44].8) [OTU(FV_FV22J.CW.[CWD.MANUAL]) ,[XIC(FV_FV22J.CW.[CWD.OUTPUT]) OTL(FV_N255[44].9) ,XIO(FV_FV22J.CW.[CWD.OUTPUT]) OTU(FV_N255[44].9) ] ] ] ,[XIC(FV_N255[44].13) OTL(FV_FV22J.CW.[CWD.CHECKOFF]) ,XIO(FV_N255[44].13) OTU(FV_FV22J.CW.[CWD.CHECKOFF]) ] ] ,XIO(Delphi_Does_Eng_Func) [[XIC(FV_FV22J.CW.[CWD.MANUAL]) OTL(FV_N255[44].8) ,XIO(FV_FV22J.CW.[CWD.MANUAL]) OTU(FV_N255[44].8) ] ,[XIC(FV_FV22J.CW.[CWD.CHECKOFF]) OTL(FV_N255[44].13) ,XIO(FV_FV22J.CW.[CWD.CHECKOFF]) OTU(FV_N255[44].13) ] ,[XIC(FV_FV22J.CW.[CWD.OUTPUT]) OTL(FV_N255[44].9) ,XIO(FV_FV22J.CW.[CWD.OUTPUT]) OTU(FV_N255[44].9) ] ] ,XIC(FV_FV22J.CW.[CWD.OUTPUT]) OTE(FV_N255[44].10) ,XIO(FV_FV22J.CW.[CWD.OUTPUT]) OTE(FV_N255[44].11) ,XIC(FV_FV22J.CW.[CWD.FAULT]) OTE(FV_N255[44].15) ];
   44: [XIC(Delphi_Does_Eng_Func) [[XIC(FV_N255[45].8) [OTL(FV_FV23C.CW.[CWD.MANUAL]) ,XIC(FV_N255[45].9) OTL(FV_FV23C.CW.[CWD.MANDRV]) ,XIO(FV_N255[45].9) OTU(FV_FV23C.CW.[CWD.MANDRV]) ] ,XIO(FV_N255[45].8) [OTU(FV_FV23C.CW.[CWD.MANUAL]) ,[XIC(FV_FV23C.CW.[CWD.OUTPUT]) OTL(FV_N255[45].9) ,XIO(FV_FV23C.CW.[CWD.OUTPUT]) OTU(FV_N255[45].9) ] ] ] ,[XIC(FV_N255[45].13) OTL(FV_FV23C.CW.[CWD.CHECKOFF]) ,XIO(FV_N255[45].13) OTU(FV_FV23C.CW.[CWD.CHECKOFF]) ] ] ,XIO(Delphi_Does_Eng_Func) [[XIC(FV_FV23C.CW.[CWD.MANUAL]) OTL(FV_N255[45].8) ,XIO(FV_FV23C.CW.[CWD.MANUAL]) OTU(FV_N255[45].8) ] ,[XIC(FV_FV23C.CW.[CWD.CHECKOFF]) OTL(FV_N255[45].13) ,XIO(FV_FV23C.CW.[CWD.CHECKOFF]) OTU(FV_N255[45].13) ] ,[XIC(FV_FV23C.CW.[CWD.OUTPUT]) OTL(FV_N255[45].9) ,XIO(FV_FV23C.CW.[CWD.OUTPUT]) OTU(FV_N255[45].9) ] ] ,XIC(FV_FV23C.CW.[CWD.OUTPUT]) OTE(FV_N255[45].10) ,XIO(FV_FV23C.CW.[CWD.OUTPUT]) OTE(FV_N255[45].11) ,XIC(FV_FV23C.CW.[CWD.FAULT]) OTE(FV_N255[45].15) ];
   45: [XIC(Delphi_Does_Eng_Func) [[XIC(FV_N255[46].8) [OTL(FV_FV23J.CW.[CWD.MANUAL]) ,XIC(FV_N255[46].9) OTL(FV_FV23J.CW.[CWD.MANDRV]) ,XIO(FV_N255[46].9) OTU(FV_FV23J.CW.[CWD.MANDRV]) ] ,XIO(FV_N255[46].8) [OTU(FV_FV23J.CW.[CWD.MANUAL]) ,[XIC(FV_FV23J.CW.[CWD.OUTPUT]) OTL(FV_N255[46].9) ,XIO(FV_FV23J.CW.[CWD.OUTPUT]) OTU(FV_N255[46].9) ] ] ] ,[XIC(FV_N255[46].13) OTL(FV_FV23J.CW.[CWD.CHECKOFF]) ,XIO(FV_N255[46].13) OTU(FV_FV23J.CW.[CWD.CHECKOFF]) ] ] ,XIO(Delphi_Does_Eng_Func) [[XIC(FV_FV23J.CW.[CWD.MANUAL]) OTL(FV_N255[46].8) ,XIO(FV_FV23J.CW.[CWD.MANUAL]) OTU(FV_N255[46].8) ] ,[XIC(FV_FV23J.CW.[CWD.CHECKOFF]) OTL(FV_N255[46].13) ,XIO(FV_FV23J.CW.[CWD.CHECKOFF]) OTU(FV_N255[46].13) ] ,[XIC(FV_FV23J.CW.[CWD.OUTPUT]) OTL(FV_N255[46].9) ,XIO(FV_FV23J.CW.[CWD.OUTPUT]) OTU(FV_N255[46].9) ] ] ,XIC(FV_FV23J.CW.[CWD.OUTPUT]) OTE(FV_N255[46].10) ,XIO(FV_FV23J.CW.[CWD.OUTPUT]) OTE(FV_N255[46].11) ,XIC(FV_FV23J.CW.[CWD.FAULT]) OTE(FV_N255[46].15) ];
   46: [XIC(Delphi_Does_Eng_Func) [[XIC(FV_N255[47].8) [OTL(FV_FV24C.CW.[CWD.MANUAL]) ,XIC(FV_N255[47].9) OTL(FV_FV24C.CW.[CWD.MANDRV]) ,XIO(FV_N255[47].9) OTU(FV_FV24C.CW.[CWD.MANDRV]) ] ,XIO(FV_N255[47].8) [OTU(FV_FV24C.CW.[CWD.MANUAL]) ,[XIC(FV_FV24C.CW.[CWD.OUTPUT]) OTL(FV_N255[47].9) ,XIO(FV_FV24C.CW.[CWD.OUTPUT]) OTU(FV_N255[47].9) ] ] ] ,[XIC(FV_N255[47].13) OTL(FV_FV24C.CW.[CWD.CHECKOFF]) ,XIO(FV_N255[47].13) OTU(FV_FV24C.CW.[CWD.CHECKOFF]) ] ] ,XIO(Delphi_Does_Eng_Func) [[XIC(FV_FV24C.CW.[CWD.MANUAL]) OTL(FV_N255[47].8) ,XIO(FV_FV24C.CW.[CWD.MANUAL]) OTU(FV_N255[47].8) ] ,[XIC(FV_FV24C.CW.[CWD.CHECKOFF]) OTL(FV_N255[47].13) ,XIO(FV_FV24C.CW.[CWD.CHECKOFF]) OTU(FV_N255[47].13) ] ,[XIC(FV_FV24C.CW.[CWD.OUTPUT]) OTL(FV_N255[47].9) ,XIO(FV_FV24C.CW.[CWD.OUTPUT]) OTU(FV_N255[47].9) ] ] ,XIC(FV_FV24C.CW.[CWD.OUTPUT]) OTE(FV_N255[47].10) ,XIO(FV_FV24C.CW.[CWD.OUTPUT]) OTE(FV_N255[47].11) ,XIC(FV_FV24C.CW.[CWD.FAULT]) OTE(FV_N255[47].15) ];
   47: [XIC(Delphi_Does_Eng_Func) [[XIC(FV_N255[48].8) [OTL(FV_FV24J.CW.[CWD.MANUAL]) ,XIC(FV_N255[48].9) OTL(FV_FV24J.CW.[CWD.MANDRV]) ,XIO(FV_N255[48].9) OTU(FV_FV24J.CW.[CWD.MANDRV]) ] ,XIO(FV_N255[48].8) [OTU(FV_FV24J.CW.[CWD.MANUAL]) ,[XIC(FV_FV24J.CW.[CWD.OUTPUT]) OTL(FV_N255[48].9) ,XIO(FV_FV24J.CW.[CWD.OUTPUT]) OTU(FV_N255[48].9) ] ] ] ,[XIC(FV_N255[48].13) OTL(FV_FV24J.CW.[CWD.CHECKOFF]) ,XIO(FV_N255[48].13) OTU(FV_FV24J.CW.[CWD.CHECKOFF]) ] ] ,XIO(Delphi_Does_Eng_Func) [[XIC(FV_FV24J.CW.[CWD.MANUAL]) OTL(FV_N255[48].8) ,XIO(FV_FV24J.CW.[CWD.MANUAL]) OTU(FV_N255[48].8) ] ,[XIC(FV_FV24J.CW.[CWD.CHECKOFF]) OTL(FV_N255[48].13) ,XIO(FV_FV24J.CW.[CWD.CHECKOFF]) OTU(FV_N255[48].13) ] ,[XIC(FV_FV24J.CW.[CWD.OUTPUT]) OTL(FV_N255[48].9) ,XIO(FV_FV24J.CW.[CWD.OUTPUT]) OTU(FV_N255[48].9) ] ] ,XIC(FV_FV24J.CW.[CWD.OUTPUT]) OTE(FV_N255[48].10) ,XIO(FV_FV24J.CW.[CWD.OUTPUT]) OTE(FV_N255[48].11) ,XIC(FV_FV24J.CW.[CWD.FAULT]) OTE(FV_N255[48].15) ];
